
                 #tempNextCmdOut.endPoint := "LKinCtrl_VecAdd"(vIn1 := #tempNextCmdIn.endPoint,
                                                               vIn2 := #tempNextCmdOut.orthogonalShiftEnd);
               ELSIF (#tempNextCmdIn.circleMode = "CM_CENTER") THEN
                 (*
                 // Calculate end point for circle mode 0 by given mode 1
                 #tempRetValue := "LKinCtrl_CalcCircEndPointWithGivenCenterAndAngle"(circleStartPoint := #tempCurrentPointRadComp,
                                                                                     circleCenterPoint := #tempNextCmdIn.circleCenterPoint,
                                                                                     pathPlane := #pathPlane,
                                                                                     pathChoice := #tempNextCmdIn.pathChoice,
                                                                                     angle := #tempNextCmdIn.circleAngle,
                                                                                     endPoint => #tempNextCmdOut.endPoint);

                 IF (#tempRetValue <> 0) THEN
                   #LKinCtrl_OffsetContour.returnValue := #tempRetValue;
                   #LKinCtrl_OffsetContour."region" := #COFF_REGION_TYPE_RAD_COMP_CIRC_NONE;
                   #LKinCtrl_OffsetContour.subBlockNumber := 35053;
                   #LKinCtrl_OffsetContour.internalNumber := 451;
                   RETURN;
                 END_IF;
                 *)
                 // Calculate end point for circle mode 0 by given mode 0
                 #tempRetValue := "LKinCtrl_CalcCircTangOrthPathPlane"(circlePoint := #tempNextCmdIn.endPoint,
                                                                       circleCenterPoint := #tempNextCmdIn.circleCenterPoint,
                                                                       pathPlane := #pathPlane,
                                                                       compDirection := #compensationDirection,
                                                                       pathChoice := #tempNextCmdIn.pathChoice,
                                                                       vUnitTangentialPathPlane => #tempNextCmdOut.tangentialUnitVecEnd,
                                                                       vUnitOrthogonalPathPlane => #tempNextCmdOut.orthogonalUnitVecEnd);

                 IF (#tempRetValue <> 0) THEN
                   #LKinCtrl_OffsetContour.returnValue := #tempRetValue;
                   #LKinCtrl_OffsetContour."region" := #COFF_REGION_TYPE_RAD_COMP_CIRC_NONE;
                   #LKinCtrl_OffsetContour.subBlockNumber := 35056;
                   #LKinCtrl_OffsetContour.internalNumber := 450;
                   RETURN;
                 END_IF;

                 // Scale othogonal vector with tool radius to get orthogonal shift
                 #tempNextCmdOut.orthogonalShiftEnd := "LKinCtrl_VecScale"(vIn := #tempNextCmdOut.orthogonalUnitVecEnd,
                                                                           factor := #toolRadius);


                 #tempNextCmdOut.endPoint := "LKinCtrl_VecAdd"(vIn1 := #tempNextCmdIn.endPoint,
                                                               vIn2 := #tempNextCmdOut.orthogonalShiftEnd);

               ELSIF (#tempNextCmdIn.circleMode = "CM_RADIUS") THEN
                 (*
                 // ------------ Via the circle radius and the end point in a main plane ("CircMode" = 2) ------------
                 // Calculate angle between center/start and center/end of circle - always the smaller one!!!
                 #tempRetValue := "LKinCtrl_CalcAngleBetweenVectors"(point1 := #tempCurrentPointRadComp,//#tempNextCmdOut.startPointOrthShifted,
                                                                     point2 := #tempNextCmdIn.endPoint,//#tempNextCmdOut.endPoint,
                                                                     intersectionPoint := #tempNextCmdIn.circleCenterPoint,
                                                                     angle => #tempAngle);

                 IF (#tempRetValue <> 0) THEN
                   #LKinCtrl_OffsetContour.returnValue := #tempRetValue;
                   #LKinCtrl_OffsetContour."region" := #COFF_REGION_TYPE_RAD_COMP_CIRC_NONE;
                   #LKinCtrl_OffsetContour.subBlockNumber := 35059;
                   #LKinCtrl_OffsetContour.internalNumber := 452;
                   RETURN;
                 END_IF;

                 // Calculate end point for circle mode 0 by given mode 2
                 #tempRetValue := "LKinCtrl_CalcCircEndPointWithGivenCenterAndAngle"(circleStartPoint := #tempCurrentPointRadComp, //tempNextCmdOut.startPointOrthShifted,
                                                                                     circleCenterPoint := #tempNextCmdIn.circleCenterPoint,
                                                                                     pathPlane := #pathPlane,
                                                                                     pathChoice := #tempNextCmdIn.pathChoice,
                                                                                     angle := #tempAngle,
                                                                                     endPoint => #tempNextCmdOut.endPoint);



                 IF (#tempRetValue <> 0) THEN
                   #LKinCtrl_OffsetContour.returnValue := #tempRetValue;
                   #LKinCtrl_OffsetContour."region" := #COFF_REGION_TYPE_RAD_COMP_CIRC_NONE;
                   #LKinCtrl_OffsetContour.subBlockNumber := 35053;
                   #LKinCtrl_OffsetContour.internalNumber := 453;
                   RETURN;
                 END_IF;
                 *)
                 ;
               END_IF;
               *)

             END_REGION
           END_IF;


           // ############# M O D I F Y   N E X T   C I R C U L A R   C O M M A N D   #############
           REGION Modify next circular command
             // Distinguish between different circular modes
             IF (#tempNextCmdIn.circleMode = "CM_BORDER") THEN

               // ------------ Via an intermediate point and the end point ("CircMode" = 0) ------------
               // Calculate intermediate point for circle mode 0 by given mode 0
               // Calculate circle paramters
               #tempRetValue := "LKinCtrl_CalcCircTangOrthPathPlane"(circlePoint :=  #tempNextCmdIn.circleIntermediatePoint,
                                                                     circleCenterPoint := #tempNextCmdIn.circleCenterPoint,
                                                                     pathPlane := #pathPlane,
                                                                     compDirection := #compensationDirection,
                                                                     pathChoice := #tempNextCmdIn.pathChoice,
                                                                     vUnitTangentialPathPlane => #tempNextCmdOut.tangentialUnitVecIntermediate,
                                                                     vUnitOrthogonalPathPlane => #tempNextCmdOut.orthogonalUnitVecIntermediate);

               IF (#tempRetValue <> 0) THEN
                 #LKinCtrl_OffsetContour.returnValue := #tempRetValue;
                 #LKinCtrl_OffsetContour."region" := #COFF_REGION_TYPE_RAD_COMP_CIRC_GEN;
                 #LKinCtrl_OffsetContour.subBlockNumber := 35056;
                 #LKinCtrl_OffsetContour.internalNumber := 460;
                 RETURN;
               END_IF;

               // Scale othogonal vector with tool radius to get orthogonal shift
               #tempNextCmdOut.orthogonalShiftIntermediate := "LKinCtrl_VecScale"(vIn := #tempNextCmdOut.orthogonalUnitVecIntermediate,
                                                                                  factor := #toolRadius);


               #tempNextCmdOut.circleIntermediatePoint := "LKinCtrl_VecAdd"(vIn1 := #tempNextCmdIn.circleIntermediatePoint,
                                                                            vIn2 := #tempNextCmdOut.orthogonalShiftIntermediate);

               // Change circle mode to 0 - intermediate point and the end point ("CircMode" = 0)
               #tempNextCmdOut.circleMode := "CM_BORDER";

             ELSIF (#tempNextCmdIn.circleMode = "CM_CENTER") THEN

               // Take care of greater angles
               #tempMod := TRUNC(#tempNextCmdIn.circleAngle / 180.0);
               IF (#tempMod >= 3) THEN
                 #tempAngle := #tempNextCmdIn.circleAngle - ((#tempMod - 1) * 180);
               ELSE
                 #tempAngle := #tempNextCmdIn.circleAngle;
               END_IF;

               // Calculate intermediate point for circle mode 0 by given mode 1
               #tempRetValue := "LKinCtrl_CalcCircEndPointWithGivenCenterAndAngle"(circleStartPoint := #tempCurrentPointRadComp, // tempNextCmdOut.startPointOrthShifted,
                                                                                   circleCenterPoint := #tempNextCmdIn.circleCenterPoint,
                                                                                   pathPlane := #pathPlane,
                                                                                   pathChoice := #tempNextCmdIn.pathChoice,
                                                                                   angle := #tempAngle / 2.0,//(#tempNextCmdIn.circleAngle / 2.0),
                                                                                   endPoint => #tempNextCmdOut.circleIntermediatePoint);
               IF (#tempRetValue <> 0) THEN
                 #LKinCtrl_OffsetContour.returnValue := #tempRetValue;
                 #LKinCtrl_OffsetContour."region" := #COFF_REGION_TYPE_RAD_COMP_CIRC_GEN;
                 #LKinCtrl_OffsetContour.subBlockNumber := 35053;
                 #LKinCtrl_OffsetContour.internalNumber := 461;
                 RETURN;
               END_IF;

               // Ceck if resulting path choice (circle with intermediate point) has changed --> circle larger than 360°
               // Calculate path choice
               #tempRetValue := "LKinCtrl_CalcCircPathChoiceByIntermediatePointAndEndPoint"(circleStartPoint := #tempCurrentPointRadComp, //tempNextCmdOut.startPointOrthShifted,
                                                                                            circleEndPoint := #tempNextCmdOut.endPoint,
                                                                                            circleintermediatePoint := #tempNextCmdOut.circleIntermediatePoint,
                                                                                            pathPlane := #pathPlane,
                                                                                            pathChoice => #tempPathChoice);


               IF (#tempRetValue <> 0) THEN
                 #LKinCtrl_OffsetContour.returnValue := #tempRetValue;
                 #LKinCtrl_OffsetContour."region" := #COFF_REGION_TYPE_RAD_COMP_CIRC_GEN;
                 #LKinCtrl_OffsetContour.subBlockNumber := 35058;
                 #LKinCtrl_OffsetContour.internalNumber := 462;
                 RETURN;
               END_IF;

               IF ((#tempNextCmdIn.pathChoice <> #tempPathChoice) OR
                 (#tempNextCmdIn.circleAngle >= 360.0))
               THEN

                 // Calculate additional angle between center/start and center/end of circle - always the smaller one!!!
                 #tempRetValue := "LKinCtrl_CalcAngleBetweenVectors"(point1 := #tempCurrentPointRadComp, //tempNextCmdOut.startPointOrthShifted,
                                                                     point2 := #tempNextCmdOut.endPoint,
                                                                     intersectionPoint := #tempNextCmdIn.circleCenterPoint,
                                                                     angle => #tempAngle);

                 IF (#tempRetValue <> 0) THEN
                   #LKinCtrl_OffsetContour.returnValue := #tempRetValue;
                   #LKinCtrl_OffsetContour."region" := #COFF_REGION_TYPE_RAD_COMP_CIRC_GEN;
                   #LKinCtrl_OffsetContour.subBlockNumber := 35059;
                   #LKinCtrl_OffsetContour.internalNumber := 463;
                   RETURN;
                 END_IF;

                 // Circle > 360° - not possible with circle type border
                 IF (#tempNextCmdIn.pathChoice <> #tempPathChoice) THEN
                   #tempNextCmdOut.circleAngle := (TRUNC((#tempNextCmdIn.circleAngle + 180.0) / 360.0) * 360.0) + #tempAngle;
                 ELSE
                   #tempNextCmdOut.circleAngle := (TRUNC((#tempNextCmdIn.circleAngle + 180.0) / 360.0) * 360.0) - #tempAngle;
                 END_IF;

                 #tempNextCmdOut.circleMode := "CM_CENTER";
               ELSE
                 // Change circle mode to 0 - intermediate point and the end point ("CircMode" = 0)
                 #tempNextCmdOut.circleMode := "CM_BORDER";
               END_IF;

             ELSIF (#tempNextCmdIn.circleMode = "CM_RADIUS") THEN
               // ------------ Via the circle radius and the end point in a main plane ("CircMode" = 2) ------------
               // Calculate angle between center/start and center/end of circle - always the smaller one!!!
               #tempRetValue := "LKinCtrl_CalcAngleBetweenVectors"(point1 := #tempCurrentPointRadComp,
                                                                   point2 := #tempNextCmdOut.endPoint,
                                                                   intersectionPoint := #tempNextCmdIn.circleCenterPoint,
                                                                   angle => #tempAngle);

               IF (#tempRetValue <> 0) THEN
                 #LKinCtrl_OffsetContour.returnValue := #tempRetValue;
                 #LKinCtrl_OffsetContour."region" := #COFF_REGION_TYPE_RAD_COMP_CIRC_GEN;
                 #LKinCtrl_OffsetContour.subBlockNumber := 35059;
                 #LKinCtrl_OffsetContour.internalNumber := 464;
                 RETURN;
               END_IF;

               // Calculate intermediate point for circle mode 0 by given mode 2
               #tempRetValue := "LKinCtrl_CalcCircEndPointWithGivenCenterAndAngle"(circleStartPoint := #tempCurrentPointRadComp, //tempNextCmdOut.startPointOrthShifted,
                                                                                   circleCenterPoint := #tempNextCmdIn.circleCenterPoint,
                                                                                   pathPlane := #pathPlane,
                                                                                   pathChoice := #tempNextCmdIn.pathChoice,
                                                                                   angle := (#tempAngle / 2.0),
                                                                                   endPoint => #tempNextCmdOut.circleIntermediatePoint);

               IF (#tempRetValue <> 0) THEN
                 #LKinCtrl_OffsetContour.returnValue := #tempRetValue;
                 #LKinCtrl_OffsetContour."region" := #COFF_REGION_TYPE_RAD_COMP_CIRC_GEN;
                 #LKinCtrl_OffsetContour.subBlockNumber := 35053;
                 #LKinCtrl_OffsetContour.internalNumber := 465;
                 RETURN;
               END_IF;

               // Change circle mode to 0 - intermediate point and the end point ("CircMode" = 0)
               #tempNextCmdOut.circleMode := "CM_BORDER";

             END_IF;

             // Additional check - has the direction between start - end and start - compensated end changed
             // --> Reversal path with "small" length (and "large" tool radius) leads to unexpected circle (mathematical correct but in an unexpected direction)
             REGION Additional plausibility check
               #tempRetValue := "LKinCtrl_CalcAngleBetweenVectors"(point1 := #tempNextCmdOut.endPoint,
                                                                   point2 := #tempNextCmdIn.endPoint,
                                                                   intersectionPoint := #tempCurrentPoint,
                                                                   angle => #tempAngle);

               IF (#tempRetValue <> 0) THEN
                 #LKinCtrl_OffsetContour.returnValue := #tempRetValue;
                 #LKinCtrl_OffsetContour."region" := #COFF_REGION_TYPE_RAD_COMP_CIRC_GEN;
                 #LKinCtrl_OffsetContour.subBlockNumber := 35059;
                 #LKinCtrl_OffsetContour.internalNumber := 470;
                 RETURN;
               END_IF;

               IF ((#tempAngle > #COFF_CIRC_REVERSAL_TOLERANCE_ANGLE) AND
                 ("LKinCtrl_VecAbs"("LKinCtrl_VecSub"(vIn1:=#tempNextCmdOut.endPoint, vIn2:=#tempNextCmdOut.circleIntermediatePoint)) < (2.0 * #toolRadius)))
               THEN
                 #LKinCtrl_OffsetContour.returnValue := #ERR_COFF_NO_SOLUTION_FOR_GIVEN_CIRCULAR_CMD;
                 #LKinCtrl_OffsetContour."region" := #COFF_REGION_TYPE_RAD_COMP_CIRC_GEN;
                 #LKinCtrl_OffsetContour.subBlockNumber := 0;
                 #LKinCtrl_OffsetContour.internalNumber := 471;
                 RETURN;
               END_IF;

             END_REGION
           END_REGION
         END_IF;
       END_REGION

     END_IF;

     // V01.00.01
     // Output before length compensation
     #pathDataOut.nextPositionAbsoluteRadComp := "LKinCtrl_3DPointToCartesianCoord"(#tempNextCmdOut.endPoint);
   END_REGION TOOL_RADIUS_COMPENSATION

   // Tool length compensation
   REGION TOOL_LENGTH_COMPENSATION
     IF (#tempToolLengthComp) THEN
       // Next command
       // -------------------------------------------------------------------------------------
       // Compensate coordinates of according to path plane
       // End point
       #tempRetValue := "LKinCtrl_CalcToolLengthCompensation"(toolLength := #toolLength,
                                                              pathPlane := #pathPlane,
                                                              point := #tempNextCmdOut.endPoint);
       IF (#tempRetValue <> 0) THEN
         #LKinCtrl_OffsetContour.returnValue := #tempRetValue;
         #LKinCtrl_OffsetContour."region" := #COFF_REGION_TYPE_LEN_COMP_NEXT;
         #LKinCtrl_OffsetContour.subBlockNumber := 35070;
         #LKinCtrl_OffsetContour.internalNumber := 601;
         RETURN;
       END_IF;

       // Circle coordinates
       IF (#tempNextCmdOut.cmdType = "LKINCTRL_MC_MOVECIRCULARABS") THEN

         IF (#tempNextCmdOut.circleMode = "CM_BORDER") THEN

           #tempRetValue := "LKinCtrl_CalcToolLengthCompensation"(toolLength := #toolLength,
                                                                  pathPlane := #pathPlane,
                                                                  point := #tempNextCmdOut.circleIntermediatePoint);
           IF (#tempRetValue <> 0) THEN
             #LKinCtrl_OffsetContour.returnValue := #tempRetValue;
             #LKinCtrl_OffsetContour."region" := #COFF_REGION_TYPE_LEN_COMP_NEXT;
             #LKinCtrl_OffsetContour.subBlockNumber := 35070;
             #LKinCtrl_OffsetContour.internalNumber := 602;
             RETURN;
           END_IF;

         ELSIF (#tempNextCmdOut.circleMode = "CM_CENTER") THEN

           #tempRetValue := "LKinCtrl_CalcToolLengthCompensation"(toolLength := #toolLength,
                                                                  pathPlane := #pathPlane,
                                                                  point := #tempNextCmdOut.circleCenterPoint);
           IF (#tempRetValue <> 0) THEN
             #LKinCtrl_OffsetContour.returnValue := #tempRetValue;
             #LKinCtrl_OffsetContour."region" := #COFF_REGION_TYPE_LEN_COMP_NEXT;
             #LKinCtrl_OffsetContour.subBlockNumber := 35070;
             #LKinCtrl_OffsetContour.internalNumber := 603;
             RETURN;
           END_IF;

         ELSIF (#tempNextCmdOut.circleMode = "CM_RADIUS") THEN
           ;
         ELSE
           #LKinCtrl_OffsetContour.returnValue := #ERR_COFF_INTERNAL; // Internal error
           #LKinCtrl_OffsetContour."region" := #COFF_REGION_TYPE_LEN_COMP_NEXT;
           #LKinCtrl_OffsetContour.internalNumber := 604;
           RETURN;
         END_IF;
       END_IF;

       // Intermediate command
       // -------------------------------------------------------------------------------------
       // Compensate coordinates of according to path plane
       IF (#tempIntermediateCmdOut.cmdType <> -1) THEN

         // End point
         #tempRetValue := "LKinCtrl_CalcToolLengthCompensation"(toolLength := #toolLength,
                                                                pathPlane := #pathPlane,
                                                                point := #tempIntermediateCmdOut.endPoint);
         IF (#tempRetValue <> 0) THEN
           #LKinCtrl_OffsetContour.returnValue := #tempRetValue;
           #LKinCtrl_OffsetContour."region" := #COFF_REGION_TYPE_LEN_COMP_INTER_CMD;
           #LKinCtrl_OffsetContour.subBlockNumber := 35070;
           #LKinCtrl_OffsetContour.internalNumber := 605;
           RETURN;
         END_IF;

         // Always circle by intemdiate point and end point
         #tempRetValue := "LKinCtrl_CalcToolLengthCompensation"(toolLength := #toolLength,
                                                                pathPlane := #pathPlane,
                                                                point := #tempIntermediateCmdOut.circleIntermediatePoint);
         IF (#tempRetValue <> 0) THEN
           #LKinCtrl_OffsetContour.returnValue := #tempRetValue;
           #LKinCtrl_OffsetContour."region" := #COFF_REGION_TYPE_LEN_COMP_INTER_CMD;
           #LKinCtrl_OffsetContour.subBlockNumber := 35070;
           #LKinCtrl_OffsetContour.internalNumber := 606;
           RETURN;
         END_IF;
       END_IF;

       // Next but one command - not needed - no output
       // -------------------------------------------------------------------------------------
      (*
       // Compensate coordinates of according to path plane
       // End point
       #tempRetValue := "LKinCtrl_CalcToolLengthCompensation"(toolLength := #toolLength,
                                                              pathPlane := #pathPlane,
                                                              point := #tempNextButOneCmdOut.endPoint);
       IF (#tempRetValue <> 0) THEN
         #LKinCtrl_OffsetContour.returnValue := #tempRetValue;
         #LKinCtrl_OffsetContour."region" := #COFF_REGION_TYPE_LEN_COMP_NEXT_BUT_ONE_CMD;
         #LKinCtrl_OffsetContour.subBlockNumber := 35070;
         #LKinCtrl_OffsetContour.internalNumber := 607
         RETURN;
       END_IF;
       *)
     END_IF;
   END_REGION

   REGION Output data

     // ############# O U T P U T   D A T A  #############
     // ###################################### 
     IF (#tempToolRadiusComp OR #tempToolLengthComp) THEN
       // Next command

       #pathDataOut.nextCommand.cmdType := #tempNextCmdOut.cmdType;
       #pathDataOut.nextCommand.cmdCoordinates.cartesianPosition := "LKinCtrl_3DPointToCartesianCoord"(#tempNextCmdOut.endPoint);

       IF (#tempNextCmdOut.cmdType = "LKINCTRL_MC_MOVECIRCULARABS") THEN
         #pathDataOut.nextCommand.cmdParameters.circleParameters.circMode := #tempNextCmdOut.circleMode;

         IF (#tempNextCmdOut.circleMode = "CM_BORDER") THEN
           #pathDataOut.nextCommand.cmdParameters.circleParameters.auxPoint[1] := #tempNextCmdOut.circleIntermediatePoint.x;
           #pathDataOut.nextCommand.cmdParameters.circleParameters.auxPoint[2] := #tempNextCmdOut.circleIntermediatePoint.y;
           #pathDataOut.nextCommand.cmdParameters.circleParameters.auxPoint[3] := #tempNextCmdOut.circleIntermediatePoint.z;

         ELSIF (#tempNextCmdOut.circleMode = "CM_CENTER") THEN
           #pathDataOut.nextCommand.cmdParameters.circleParameters.pathChoice := #tempNextCmdIn.pathChoice;
           #pathDataOut.nextCommand.cmdParameters.circleParameters.circlePlane := #tempNextCmdIn.circlePlane;
           #pathDataOut.nextCommand.cmdParameters.circleParameters.auxPoint[1] := #tempNextCmdOut.circleCenterPoint.x;
           #pathDataOut.nextCommand.cmdParameters.circleParameters.auxPoint[2] := #tempNextCmdOut.circleCenterPoint.y;
           #pathDataOut.nextCommand.cmdParameters.circleParameters.auxPoint[3] := #tempNextCmdOut.circleCenterPoint.z;
           #pathDataOut.nextCommand.cmdParameters.circleParameters.arc := #tempNextCmdOut.circleAngle; // #tempNextCmdIn.circleAngle;

         ELSIF (#tempNextCmdOut.circleMode = "CM_RADIUS") THEN
           #pathDataOut.nextCommand.cmdParameters.circleParameters.pathChoice := #tempNextCmdIn.pathChoice;
           #pathDataOut.nextCommand.cmdParameters.circleParameters.circlePlane := #tempNextCmdIn.circlePlane;
           #pathDataOut.nextCommand.cmdParameters.circleParameters.radius := #tempNextCmdIn.circleRadius;

         ELSE
           #LKinCtrl_OffsetContour.returnValue := #ERR_COFF_INTERNAL; // Internal error
           #LKinCtrl_OffsetContour."region" := #COFF_REGION_TYPE_OUTPUT_DATA;
           RETURN;
         END_IF;
       END_IF;

       // Coordinate a
       // ------------
       // Linear absolute
       IF (#tempNextCmdIn.cmdType = "LKINCTRL_MC_MOVELINEARABS") THEN
         // Absolute coordinates
         #pathDataOut.nextCommand.cmdCoordinates.cartesianPosition.a := #pathDataIn.nextCommand.cmdCoordinates.cartesianPosition.a;
         // Linear relative
       ELSIF (#tempNextCmdIn.cmdType = "LKINCTRL_MC_MOVELINEARREL") THEN
         // Relative coordinates -> calculate absolute coordinate (always)
         #pathDataOut.nextCommand.cmdCoordinates.cartesianPosition.a := #pathDataIn.currentPos.positionAbsolute.a + #pathDataIn.nextCommand.cmdCoordinates.cartesianPosition.a;
         // Circular absolute  
       ELSIF (#tempNextCmdIn.cmdType = "LKINCTRL_MC_MOVECIRCULARABS") THEN
         // Absolute coordinates
         #pathDataOut.nextCommand.cmdCoordinates.cartesianPosition.a := #pathDataIn.nextCommand.cmdCoordinates.cartesianPosition.a;
         // Circular relative  
       ELSIF (#tempNextCmdIn.cmdType = "LKINCTRL_MC_MOVECIRCULARREL") THEN
         // Relative coordinates -> calculate absolute coordinate (always)
         #pathDataOut.nextCommand.cmdCoordinates.cartesianPosition.a := #pathDataIn.currentPos.positionAbsolute.a + #pathDataIn.nextCommand.cmdCoordinates.cartesianPosition.a;
       END_IF;

       // Output absolute end point for next cycle (including coordinate a)
       #pathDataOut.nextPositionAbsolute := "LKinCtrl_3DPointToCartesianCoord"(#tempNextCmdIn.endPoint);
       #pathDataOut.nextPositionAbsolute.a := #pathDataOut.nextCommand.cmdCoordinates.cartesianPosition.a;

       // Output absolute end point (radius compensated) for next cycle (including coordinate a)
       // V01.00.01
       // #pathDataOut.nextPositionAbsoluteRadComp := "LKinCtrl_3DPointToCartesianCoord"(#tempNextCmdOut.endPoint);
       #pathDataOut.nextPositionAbsoluteRadComp.a := #pathDataOut.nextCommand.cmdCoordinates.cartesianPosition.a;

       // Intermediate command
       IF (#tempIntermediateCmdOut.cmdType <> -1) THEN

         // Take all parameter preliminary
         #pathDataOut.intermediateCommand := #pathDataIn.nextCommand;

         #pathDataOut.intermediateCommand.cmdType := #tempIntermediateCmdOut.cmdType;
         #pathDataOut.intermediateCommand.cmdParameters.circleParameters.circMode := #tempIntermediateCmdOut.circleMode;

         // Circle by intemdiate point and end point
         #pathDataOut.intermediateCommand.cmdCoordinates.cartesianPosition := "LKinCtrl_3DPointToCartesianCoord"(#tempIntermediateCmdOut.endPoint);
         #pathDataOut.intermediateCommand.cmdParameters.circleParameters.auxPoint[1] := #tempIntermediateCmdOut.circleIntermediatePoint.x;
         #pathDataOut.intermediateCommand.cmdParameters.circleParameters.auxPoint[2] := #tempIntermediateCmdOut.circleIntermediatePoint.y;
         #pathDataOut.intermediateCommand.cmdParameters.circleParameters.auxPoint[3] := #tempIntermediateCmdOut.circleIntermediatePoint.z;

         // Coordinate a
         #pathDataOut.intermediateCommand.cmdCoordinates.cartesianPosition.a := #pathDataOut.nextCommand.cmdCoordinates.cartesianPosition.a;
       ELSE
         #pathDataOut.intermediateCommand.cmdType := -1;
       END_IF;

       // Next but one command
       //#pathDataOut.nextButOneCommand.cmdType := #tempNextButOneCmdIn.cmdType;
       //#pathDataOut.nextButOneCommand.cmdCoordinates.cartesianPosition := "LKinCtrl_3DPointToCartesianCoord"(#tempNextButOneCmdOut.endPoint);
       #pathDataOut.nextButOneCommand.transitionParameter[1] := #tempNextButOneCmdOut.transitionParameter1;
     ELSE
       // Next command
       #pathDataOut.nextCommand := #pathDataIn.nextCommand;
     END_IF;

   END_REGION

   #LKinCtrl_OffsetContour.returnValue := 16#0;
   #LKinCtrl_OffsetContour."region" := #COFF_REGION_TYPE_NONE;
   #LKinCtrl_OffsetContour.subBlockNumber := 16#0;
   #LKinCtrl_OffsetContour.internalNumber := 0;
END_FUNCTION

// folder: LKinCtrl_Blocks/LKinCtrl_SubBlocks/LKinCtrl_ContOffsetBlocks/LKinCtrl_ContOffset_SubBlocks

FUNCTION "LKinCtrl_CheckInnerOuterCorner" : Word   // FC35051, SCL
TITLE = LKinCtrl_CheckInnerOuterCorner
{ S7_Optimized_Access := 'TRUE' }
AUTHOR : tech.team.motioncontrol@siemens.com
FAMILY : LKinCtrl
VERSION : 1.1
// Check for inner or outer corner
   VAR_INPUT
      vInFirst : "LKinCtrl_typeCOff3DPoint";   // Input vector first
      vInSecond : "LKinCtrl_typeCOff3DPoint";   // Input vector second
      pathPlane : Int;   // Path plane: XZ= 0, YZ=1, XY= 2
      direction : Int;   // Tool radius compensation direction: left=1, right = 0
   END_VAR
   VAR_OUTPUT
      cornerType : Int;   // Corner type - 0: outer corner, 1: inner corner
   END_VAR
   VAR_TEMP
      tempCrossVec : "LKinCtrl_typeCOff3DPoint";
   END_VAR
   // Ret_Val : Return value
   VAR CONSTANT
      ERR_COFF_INVALID_PATH_PLANE : Word := 16#8303;   // Invalid path plane
      ERR_COFF_INVALID_COMPENSATION_DIRECTION : Word := 16#8304;   // Invalid compensation direction
   END_VAR
BEGIN
   //=============================================================================
   // SIEMENS AG
   // (c)Copyright 2019 All Rights Reserved
   //-----------------------------------------------------------------------------
   // Library: - 
   // Tested with: S7-1516T-3 PN
   // Engineering: TIA Portal V15
   // Restrictions: -
   // Requirements: S7-1500/S7-1500T FW 2.5
   // Functionality: Check for inner or outer corner
   //-----------------------------------------------------------------------------
   // Change log table:
   // Version  Date       Expert in charge Changes applied
   // 01.00.00 2019-01-24 AW               created
   // 01.00.01 2020-10-13 AW               bugfix - path plane CP_XZ - different orientation, not against third axis!
   //=============================================================================
   REGION PLAUSIBILITY_CHECK
     // Check path plane
     IF ((#pathPlane >= "CP_XZ") AND (#pathPlane <= "CP_XY"))
     THEN
       // Check compensation direction
       IF ((#direction >= "LKINCTRL_COMP_LEFT") AND (#direction <= "LKINCTRL_COMP_RIGHT"))
       THEN
         ;
       ELSE
         #LKinCtrl_CheckInnerOuterCorner := #ERR_COFF_INVALID_COMPENSATION_DIRECTION; // Invalid compensation direction
         RETURN;
       END_IF;
     ELSE
       #LKinCtrl_CheckInnerOuterCorner := #ERR_COFF_INVALID_PATH_PLANE; // Invalid path plane
       RETURN;
     END_IF;
   END_REGION PLAUSIBILITY_CHECK

   REGION CALCULATION
     #tempCrossVec := "LKinCtrl_VecCrossProd"(vIn1 := #vInFirst,
                                              vIn2 := #vInSecond);

   // Check path plane
   IF (#pathPlane = "CP_XY") THEN
     IF (#direction = "LKINCTRL_COMP_RIGHT") THEN
       IF (#tempCrossVec.z > 0.0) THEN
         #cornerType := "LKINCTRL_OUTER_CORNER";
       ELSE
         #cornerType := "LKINCTRL_INNER_CORNER";
       END_IF;
     ELSE
       IF (#tempCrossVec.z < 0.0) THEN
         #cornerType := "LKINCTRL_OUTER_CORNER";
       ELSE
         #cornerType := "LKINCTRL_INNER_CORNER";
       END_IF;
     END_IF;

   // 2020-10-13 AW path plane CP_XZ - different orientation, not against third axis!
   // direction changed
   ELSIF (#pathPlane = "CP_XZ") THEN
       IF (#direction = "LKINCTRL_COMP_RIGHT") THEN
         IF (#tempCrossVec.y > 0.0) THEN
           #cornerType := "LKINCTRL_INNER_CORNER";
         ELSE
           #cornerType := "LKINCTRL_OUTER_CORNER";
         END_IF;
       ELSE
         IF (#tempCrossVec.y < 0.0) THEN
           #cornerType := "LKINCTRL_INNER_CORNER";
         ELSE
           #cornerType := "LKINCTRL_OUTER_CORNER";
         END_IF;
       END_IF;
     ELSIF (#pathPlane = "CP_YZ") THEN
     IF (#direction = "LKINCTRL_COMP_RIGHT") THEN
       IF (#tempCrossVec.x > 0.0) THEN
         #cornerType := "LKINCTRL_OUTER_CORNER";
       ELSE
         #cornerType := "LKINCTRL_INNER_CORNER";
       END_IF;
     ELSE
       IF (#tempCrossVec.x < 0.0) THEN
         #cornerType := "LKINCTRL_OUTER_CORNER";
       ELSE
         #cornerType := "LKINCTRL_INNER_CORNER";
       END_IF;
     END_IF;
   END_IF;

   #LKinCtrl_CheckInnerOuterCorner := 0;
   END_REGION CALCULATION
END_FUNCTION

FUNCTION "LKinCtrl_CalcCircCenterByRadiusAndEndPoint" : Word   // FC35052, SCL
TITLE = LKinCtrl_CalcCircCenterByRadiusAndEndPoint
{ S7_Optimized_Access := 'TRUE' }
AUTHOR : tech.team.motioncontrol@siemens.com
FAMILY : LKinCtrl
VERSION : 1.0
// Calculate circle center point with given start point, end point and radius
   VAR_INPUT
      circleStartPoint : "LKinCtrl_typeCOff3DPoint";   // Circle start point
      circleEndPoint : "LKinCtrl_typeCOff3DPoint";   // Circle end point
      pathPlane : Int;   // Path plane: XZ= 0, YZ=1, XY= 2
      circleRadius : LReal;   // Circle radius
      pathChoice : DInt;   // Circle path choice: positive= 0, negative= 1
   END_VAR
   VAR_OUTPUT
      circCenterPoint : "LKinCtrl_typeCOff3DPoint";   // Circle center point
   END_VAR
   VAR_TEMP
      tempRetValue : Word;
      tempPa : "LKinCtrl_typeCOff3DPoint";
      tempPb : "LKinCtrl_typeCOff3DPoint";
      tempVEndStart : "LKinCtrl_typeCOff3DPoint";
      tempVPaStart : "LKinCtrl_typeCOff3DPoint";
      tempCrossVec : "LKinCtrl_typeCOff3DPoint";
   END_VAR
   // Ret_Val : Return value
   VAR CONSTANT
      ERR_COFF_INVALID_PATH_PLANE : Word := 16#8303;   // Error - invalid path plane
   END_VAR
BEGIN
   //=============================================================================
   // SIEMENS AG
   // (c)Copyright 2019 All Rights Reserved
   //-----------------------------------------------------------------------------
   // Library: - 
   // Tested with: S7-1516T-3 PN
   // Engineering: TIA Portal V15
   // Restrictions: -
   // Requirements: S7-1500/S7-1500T FW 2.5
   // Functionality: Calculate circle center point with given start point, end point and radius
   //-----------------------------------------------------------------------------
   // Change log table:
   // Version  Date       Expert in charge Changes applied
   // 01.00.00 2019-01-24 AW               created
   //=============================================================================

   REGION PLAUSIBILITY_CHECK
     // Check path plane
     IF ((#pathPlane >= "CP_XZ") AND (#pathPlane <= "CP_XY"))
     THEN
       ;
     ELSE
       #LKinCtrl_CalcCircCenterByRadiusAndEndPoint := #ERR_COFF_INVALID_PATH_PLANE; // Invalid path plane
       RETURN;
     END_IF;
   END_REGION PLAUSIBILITY_CHECK

   REGION CALCULATION


     // Calculate circle center point by letting the following two circles intersect
     // 1st circle around start point with radius
     // 2nd circle around end point with radius
     #tempRetValue := "LKinCtrl_CalcCircleCircleIntersectionPoint"(circleCenterPoint1 := #circleStartPoint,
                                                                   circleCenterPoint2 := #circleEndPoint,
                                                                   circleRadius1 := #circleRadius,
                                                                   circleRadius2 := #circleRadius,
                                                                   pathPlane := #pathPlane,
                                                                   intersectionPointA => #tempPa,
                                                                   intersectionPointB => #tempPb);

     IF (#tempRetValue <> 16#0) THEN
       #LKinCtrl_CalcCircCenterByRadiusAndEndPoint := #tempRetValue;
       RETURN;
     END_IF;

     // Which one ist the correct circle center point? Calculate left and right

     // Difference vectors
     #tempVEndStart := "LKinCtrl_VecSub"(vIn1 := #circleEndPoint, vIn2 := #circleStartPoint);
     #tempVPaStart := "LKinCtrl_VecSub"(vIn1 := #tempPa, vIn2 := #circleStartPoint);
     #tempCrossVec := "LKinCtrl_VecCrossProd"(vIn1 := #tempVEndStart,
                                              vIn2 := #tempVPaStart);

     // Check path plane
     IF (#pathPlane = "CP_XY") THEN
       IF (#tempCrossVec.z > 0.0) THEN
         IF (#pathChoice = 0) THEN
           #circCenterPoint := #tempPa;
         ELSE
           #circCenterPoint := #tempPb;
         END_IF;
       ELSE
         // Todo - is the else necessary?
         IF (#pathChoice = 0) THEN
           #circCenterPoint := #tempPb;
         ELSE
           #circCenterPoint := #tempPa;
         END_IF;
       END_IF;
     ELSIF (#pathPlane = "CP_XZ") THEN
       IF (#tempCrossVec.y > 0.0) THEN
         IF (#pathChoice = 0) THEN
           #circCenterPoint := #tempPa;
         ELSE
           #circCenterPoint := #tempPb;
         END_IF;
       ELSE
         IF (#pathChoice = 0) THEN
           #circCenterPoint := #tempPb;
         ELSE
           #circCenterPoint := #tempPa;
         END_IF;
       END_IF;
     ELSIF (#pathPlane = "CP_YZ") THEN
       IF (#tempCrossVec.x > 0.0) THEN
         IF (#pathChoice = 0) THEN
           #circCenterPoint := #tempPa;
         ELSE
           #circCenterPoint := #tempPb;
         END_IF;
       ELSE
         IF (#pathChoice = 0) THEN
           #circCenterPoint := #tempPb;
         ELSE
           #circCenterPoint := #tempPa;
         END_IF;
       END_IF;
     END_IF;

   END_REGION ; 
   #LKinCtrl_CalcCircCenterByRadiusAndEndPoint := 0; // o.k.
END_FUNCTION

FUNCTION "LKinCtrl_CalcCircEndPointWithGivenCenterAndAngle" : Word   // FC35053, SCL
TITLE = LKinCtrl_CalcCircEndPointWithGivenCenterAndAngle
{ S7_Optimized_Access := 'TRUE' }
AUTHOR : tech.team.motioncontrol@siemens.com
FAMILY : LKinCtrl
VERSION : 1.0
// Calculate circle end point with given start point, circle center and angle
   VAR_INPUT
      circleStartPoint : "LKinCtrl_typeCOff3DPoint";   // Circle start point
      circleCenterPoint : "LKinCtrl_typeCOff3DPoint";   // Circle center point
      pathPlane : Int;   // Path plane: XZ= 0, YZ=1, XY= 2
      pathChoice : DInt;   // Circle path choice: positive= 0, negative= 1
      angle : LReal;   // Circle angle
   END_VAR
   VAR_OUTPUT
      endPoint : "LKinCtrl_typeCOff3DPoint";
   END_VAR
   VAR_TEMP
      tempSin : LReal;
      tempCos : LReal;
      tempVOrthogonal : "LKinCtrl_typeCOff3DPoint";   // Othogonal vector
      tempVRotated : "LKinCtrl_typeCOff3DPoint";
   END_VAR
   VAR CONSTANT
      ERR_COFF_INVALID_PATH_PLANE : Word := 16#8303;   // Error - invalid path plane
      ERR_COFF_INVALID_COMPENSATION_DIRECTION : Word := 16#8304;   // Error - invalid compensation direction
   END_VAR
BEGIN
   //=============================================================================
   // SIEMENS AG
   // (c)Copyright 2019 All Rights Reserved
   //-----------------------------------------------------------------------------
   // Library: - 
   // Tested with: S7-1516T-3 PN
   // Engineering: TIA Portal V15
   // Restrictions: -
   // Requirements: S7-1500/S7-1500T FW 2.5
   // Functionality: Calculate circle end point with given
   // start point, circle center and angle
   //-----------------------------------------------------------------------------
   // Change log table:
   // Version  Date       Expert in charge Changes applied
   // 01.00.00 2019-01-24 AW               created
   //=============================================================================

   REGION PLAUSIBILITY_CHECK
     // Check path plane
     IF ((#pathPlane >= "CP_XZ") AND (#pathPlane <= "CP_XY"))
     THEN
       // Check compensation direction
       IF ((#pathChoice >= 0) AND (#pathChoice <= 1))
       THEN
         ;
       ELSE
         #LKinCtrl_CalcCircEndPointWithGivenCenterAndAngle := #ERR_COFF_INVALID_COMPENSATION_DIRECTION; // Invalid compensation direction
         RETURN;
       END_IF;
     ELSE
       #LKinCtrl_CalcCircEndPointWithGivenCenterAndAngle := #ERR_COFF_INVALID_PATH_PLANE; // Invalid path plane
       RETURN;
     END_IF;
   END_REGION PLAUSIBILITY_CHECK

   REGION CALCULATION

   // Calc radius vector (difference vector) circle center to start point
   #tempVOrthogonal := "LKinCtrl_VecSub"(vIn1 := #circleStartPoint, vIn2 := #circleCenterPoint);

   IF (#pathChoice = 0) THEN
     // positive
     #tempSin := SIN(#angle * "LKINCTRL_PI" / 180.0);
     #tempCos := COS(#angle * "LKINCTRL_PI" / 180.0);
   ELSE
     #tempSin := SIN(- #angle * "LKINCTRL_PI" / 180.0);
     #tempCos := COS(- #angle * "LKINCTRL_PI" / 180.0);
   END_IF;

   // Check path plane
   IF (#pathPlane = "CP_XY") THEN
     // Rotation around Z
     #tempVRotated.x := #tempVOrthogonal.x * #tempCos - #tempVOrthogonal.y * #tempSin;      // Calculation X
     #tempVRotated.y := #tempVOrthogonal.x * #tempSin + #tempVOrthogonal.y * #tempCos;      // Calculation Y
     #tempVRotated.z := #tempVOrthogonal.z;                                                 // Calculation Z

   ELSIF (#pathPlane = "CP_XZ") THEN
     // Rotation around Y
     #tempVRotated.x := #tempVOrthogonal.x * #tempCos + #tempVOrthogonal.z * #tempSin;      // Calculation X
     #tempVRotated.y := #tempVOrthogonal.y;                                                 // Calculation Y
     #tempVRotated.z := -#tempVOrthogonal.x * #tempSin + #tempVOrthogonal.z * #tempCos;     // Calculation Z

   ELSIF (#pathPlane = "CP_YZ") THEN
     // Rotation around X
     #tempVRotated.x := #tempVOrthogonal.x;      // Calculation X
     #tempVRotated.y := #tempVOrthogonal.y * #tempCos - #tempVOrthogonal.z * #tempSin;       // Calculation Y
     #tempVRotated.z := #tempVOrthogonal.y * #tempSin + #tempVOrthogonal.z * #tempCos;     // Calculation Z
   END_IF;

   // Calculate end point of circle by adding the rotated vector to the circle center point
   #endPoint := "LKinCtrl_VecAdd"(vIn1:=#tempVRotated, vIn2:=#circleCenterPoint);

   END_REGION CALCULATION

   #LKinCtrl_CalcCircEndPointWithGivenCenterAndAngle := 0;
END_FUNCTION

FUNCTION "LKinCtrl_CalcCircleIntermediatePos" : Void   // FC35054, SCL
TITLE = LKinCtrl_CalcCircleIntermediatePos
{ S7_Optimized_Access := 'TRUE' }
AUTHOR : tech.team.motioncontrol@siemens.com
FAMILY : LKinCtrl
VERSION : 1.0
// Calculate intermediate point of circle with given initial end point, calculated end point and tool radius
   VAR_INPUT
      initialEndPoint : "LKinCtrl_typeCOff3DPoint";   // Initial end point
      newEndPoint : "LKinCtrl_typeCOff3DPoint";   // New calculated end point
      toolRadius : LReal;   // Tool radius
   END_VAR
   VAR_OUTPUT
      circIntermediatePoint : "LKinCtrl_typeCOff3DPoint";   // circle intermediate point
   END_VAR
   VAR_TEMP
      tempVecDiff : "LKinCtrl_typeCOff3DPoint";
      tempUnitVecDiff : "LKinCtrl_typeCOff3DPoint";
   END_VAR
BEGIN
   //=============================================================================
   // SIEMENS AG
   // (c)Copyright 2019 All Rights Reserved
   //-----------------------------------------------------------------------------
   // Library: - 
   // Tested with: S7-1516T-3 PN
   // Engineering: TIA Portal V15
   // Restrictions: -
   // Requirements: S7-1500/S7-1500T FW 2.5
   // Functionality: Calculate intermediate point of circle
   // with given initial end point, calculated end point and tool radius
   //-----------------------------------------------------------------------------
   // Change log table:
   // Version  Date       Expert in charge Changes applied
   // 01.00.00 2019-02-05 AW               created
   //=============================================================================

   REGION PLAUSIBILITY_CHECK
   END_REGION PLAUSIBILITY_CHECK

   REGION CALCULATION
   // Difference vector between new end point and initial end point
   #tempVecDiff := "LKinCtrl_VecSub"(vIn1 := #newEndPoint,
                                  vIn2 := #initialEndPoint);

   // Calculate direction vetor to intermediate point
   #tempUnitVecDiff := "LKinCtrl_VecUnit"(#tempVecDiff);

   // Calculate intermediate point: initialEndPoint + lambda * radius
   #circIntermediatePoint := "LKinCtrl_VecAdd"(vIn1:= #initialEndPoint, vIn2:= "LKinCtrl_VecScale"(vIn := #tempUnitVecDiff, factor := #toolRadius));

   END_REGION CALCULATION
END_FUNCTION

FUNCTION "LKinCtrl_CalcLineTangOrthPathPlane" : Word   // FC35055, SCL
TITLE = LKinCtrl_CalcLineTangOrthPathPlane
{ S7_Optimized_Access := 'TRUE' }
AUTHOR : tech.team.motioncontrol@siemens.com
FAMILY : LKinCtrl
VERSION : 1.0
// Calculate orthogonal and tangential vector of a line with respect ot the path plane
   VAR_INPUT
      pathPlane : Int;   // Path plane: XZ= 0, YZ=1, XY= 2
      compDirection : Int;   // Tool radius compensation direction: left=1, right = 0
      vInFirst : "LKinCtrl_typeCOff3DPoint";   // Next position
      vInSecond : "LKinCtrl_typeCOff3DPoint";   // Current position
   END_VAR
   VAR_OUTPUT
      vUnitTangentialPathPlane : "LKinCtrl_typeCOff3DPoint";   // Output tangential vector - path plane - unit vector
      vUnitOrthogonalPathPlane : "LKinCtrl_typeCOff3DPoint";   // Output orthogonal vector - path plane - unit vector
   END_VAR
   VAR_TEMP
      tempVOrthogonal : "LKinCtrl_typeCOff3DPoint";   // Othogonal vector
      tempVTangential : "LKinCtrl_typeCOff3DPoint";   // Tangential vector
   END_VAR
   VAR CONSTANT
      ERR_COFF_INVALID_PATH_PLANE : Word := 16#8303;   // Error - invalid path plane
      ERR_COFF_INVALID_COMPENSATION_DIRECTION : Word := 16#8304;   // Error - invalid compensation direction
   END_VAR
BEGIN
   //=============================================================================
   // SIEMENS AG
   // (c)Copyright 2019 All Rights Reserved
   //-----------------------------------------------------------------------------
   // Library: - 
   // Tested with: S7-1516T-3 PN
   // Engineering: TIA Portal V15
   // Restrictions: -
   // Requirements: S7-1500/S7-1500T FW 2.5
   // Functionality: Calculate orthogonal and tangential vector of a line
   // with respect ot the path plane
   //-----------------------------------------------------------------------------
   // Change log table:
   // Version  Date       Expert in charge Changes applied
   // 01.00.00 2019-02-05 AW               created
   //=============================================================================

   REGION PLAUSIBILITY_CHECK
   // Check path plane
     IF ((#pathPlane >= "CP_XZ") AND (#pathPlane <= "CP_XY"))
   THEN
     // Check compensation direction
     IF ((#compDirection >= "LKINCTRL_COMP_LEFT") AND (#compDirection <= "LKINCTRL_COMP_RIGHT"))
     THEN
       ;
     ELSE
       #LKinCtrl_CalcLineTangOrthPathPlane := #ERR_COFF_INVALID_COMPENSATION_DIRECTION; // Invalid compensation direction
       RETURN;
     END_IF;
   ELSE
     #LKinCtrl_CalcLineTangOrthPathPlane := #ERR_COFF_INVALID_PATH_PLANE; // Invalid path plane
     RETURN;
   END_IF;

   END_REGION PLAUSIBILITY_CHECK

   REGION CALCULATION
     // Calculate difference vector (take care of path plane) - tangential vector
     #tempVTangential := "LKinCtrl_VecSub"(vIn1 := #vInFirst,
                                           vIn2 := #vInSecond);

     // Take care of path plane
     CASE #pathPlane OF
       "CP_XY":
         #tempVTangential.z := 0.0;

       "CP_XZ":
         #tempVTangential.y := 0.0;

       "CP_YZ":
         #tempVTangential.x := 0.0;
     END_CASE;

     // Normalize vector
     #tempVTangential := "LKinCtrl_VecUnit"(vIn := #tempVTangential);


   // Calculate orthogonal vector to current vector depending on path plane and compensation direction
   CASE #pathPlane OF
     "CP_XY":
       IF (#compDirection = "LKINCTRL_COMP_LEFT") THEN
         #tempVOrthogonal.x := - #tempVTangential.y;
         #tempVOrthogonal.y := #tempVTangential.x;
         #tempVOrthogonal.z := 0.0;
       ELSE
         #tempVOrthogonal.x := #tempVTangential.y;
         #tempVOrthogonal.y := - #tempVTangential.x;
         #tempVOrthogonal.z := 0.0;          
       END_IF;

     "CP_XZ":
       (*
       IF (#compDirection = "LKINCTRL_COMP_LEFT") THEN
         #tempVOrthogonal.x := #tempVTangential.z;
         #tempVOrthogonal.y := 0.0;
         #tempVOrthogonal.z := - #tempVTangential.x;
       ELSE
         #tempVOrthogonal.x := - #tempVTangential.z;
         #tempVOrthogonal.y := 0.0;
         #tempVOrthogonal.z := #tempVTangential.x;
       END_IF;*)

       IF (#compDirection = "LKINCTRL_COMP_LEFT") THEN
         #tempVOrthogonal.x := -#tempVTangential.z;
         #tempVOrthogonal.y := 0.0;
         #tempVOrthogonal.z := #tempVTangential.x;
       ELSE
         #tempVOrthogonal.x := #tempVTangential.z;
         #tempVOrthogonal.y := 0.0;
         #tempVOrthogonal.z := -#tempVTangential.x;
       END_IF;

